REGION Network 15: DB62.DBX7.6 = Soot System Opacity
   // Word 4 bit 14
   RUNG wire#powerrail
      I_Contact( "10 DI_DATA".E700_OPACITY )
      { S7_Templates := "SrcType := Int" } GE_Contact(in1 := "100_BC_AUTO_SEQ_DB".CRNT_STEP, in2 := 240)
      Coil( %DB62.DBX7.6 )
   END_RUNG
   // the same network as SCL:
   %DB62.DBX7.6 := NOT "10 DI_DATA".E700_OPACITY AND ("100_BC_AUTO_SEQ_DB".CRNT_STEP >= 240);
END_REGION

REGION Network 16: DB62.DBX7.7 = Soot System Out of Range
   // Word 4 bit 15
   RUNG wire#powerrail
      "IDB_E700 Alarms"(Value := "12_AI_Data".E700SootContentIn, "Raw Value" := "IG Soot Content", Enable := true, "SHORT CIRCUIT VALUE" := 32000.0, "BROKEN WIRE VALUE" := -32000.0, "VERY LOW LEVEL VALUE (LL)" :=, "LOW LEVEL VALUE (L)" :=, "HIGH LEVEL VALUE (H)" :=, "VERY HIGH LEVEL VALUE (HH)" :=, OFFSET :=, "ALARM DELAY" :=, "Peak Value Reset" :=, "ALARM HH" =>, "ALARM H" =>, "ALARM L" =>, "ALARM LL" =>, "ALARM READING" => %DB62.DBX7.7, "Peak Value" =>, Alarm =>, Alarm_INT =>, "Enable Delay Time" :=, "High Value Release" :=)
   END_RUNG
   // the same network as SCL:
   "IDB_E700 Alarms"(Value := "12_AI_Data".E700SootContentIn,   // "502_ALM_ANALOG"
                     "Raw Value" := "IG Soot Content",
                     Enable := true,
                     "SHORT CIRCUIT VALUE" := 32000.0,
                     "BROKEN WIRE VALUE" := -32000.0,
                     "ALARM READING" => %DB62.DBX7.7);
END_REGION

REGION Network 17: DB62.DBX4.6 = E131 I&A Compresor Warning
   // Word 3 bit 6
   RUNG wire#powerrail
      I_Contact( "10 DI_DATA".E131_WRNG )
      Coil( %DB62.DBX4.6 )
   END_RUNG
   // the same network as SCL:
   %DB62.DBX4.6 := NOT "10 DI_DATA".E131_WRNG;
END_REGION

REGION Network 18: DB62.DBX4.7 = E131 I&A Compresor Not Running
   // Word 3 bit 7          Supresed. Not Available on The Bordeira
   RUNG wire#powerrail
      I_Contact( "10 DI_DATA".E131_OK )
      { S7_Templates := "SrcType := Int" } GT_Contact(in1 := "100_BC_AUTO_SEQ_DB".CRNT_STEP, in2 := 1)
      Contact( "AlwaysFALSE" )
      Coil( %DB62.DBX4.7 )
   END_RUNG
   // the same network as SCL:
   %DB62.DBX4.7 := NOT "10 DI_DATA".E131_OK AND ("100_BC_AUTO_SEQ_DB".CRNT_STEP > 1) AND "AlwaysFALSE";
END_REGION

REGION Network 19: DB62.DBX_ =IW98 - Flame Signal (FD-001)
   // Word 1 bit 12
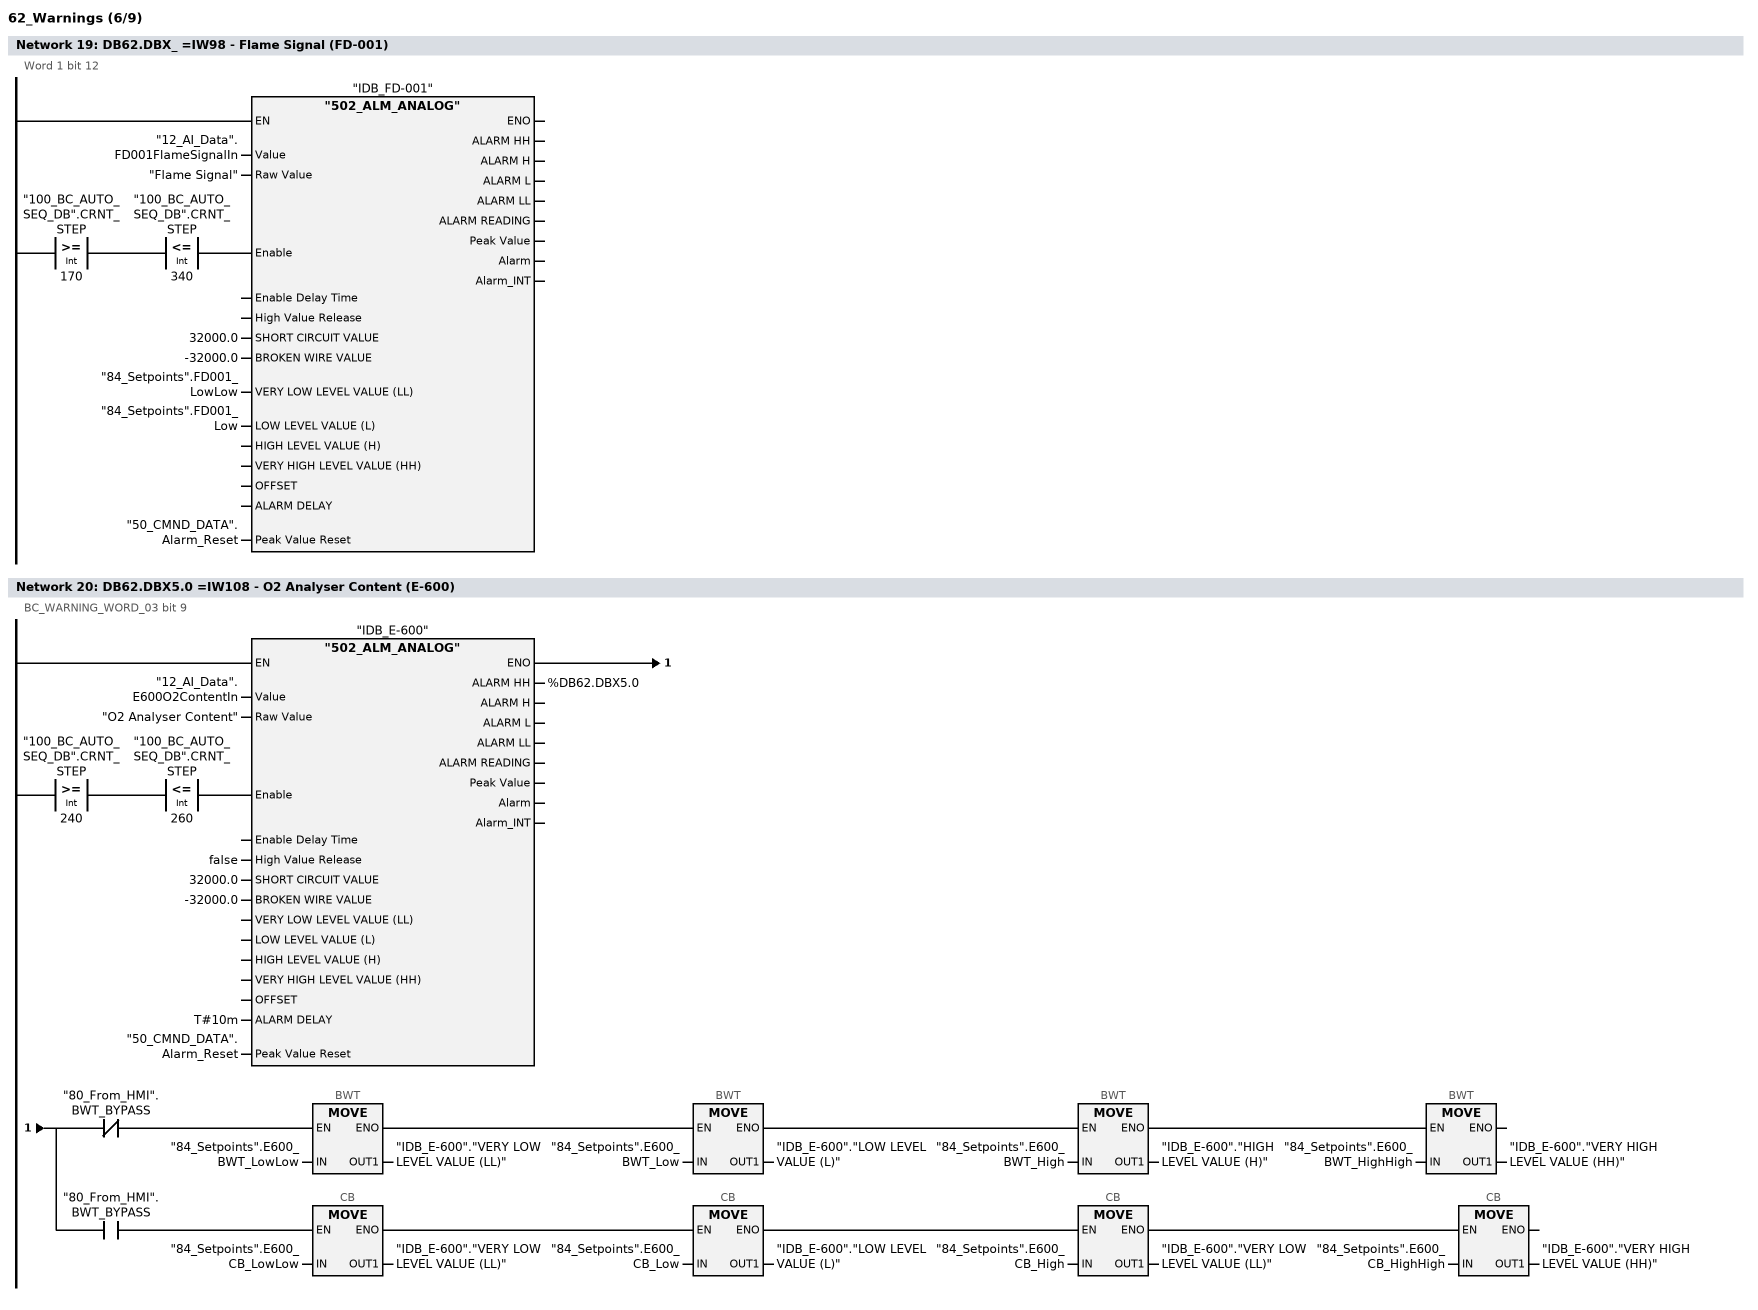
   RUNG wire#powerrail
      "IDB_FD-001"(Enable := wire#w1, Value := "12_AI_Data".FD001FlameSignalIn, "Raw Value" := "Flame Signal", "SHORT CIRCUIT VALUE" := 32000.0, "BROKEN WIRE VALUE" := -32000.0, "VERY LOW LEVEL VALUE (LL)" := "84_Setpoints".FD001_LowLow, "LOW LEVEL VALUE (L)" := "84_Setpoints".FD001_Low, "HIGH LEVEL VALUE (H)" :=, "VERY HIGH LEVEL VALUE (HH)" :=, OFFSET :=, "ALARM DELAY" :=, "Peak Value Reset" := "50_CMND_DATA".Alarm_Reset, "ALARM HH" =>, "ALARM H" =>, "ALARM L" =>, "ALARM LL" =>, "ALARM READING" =>, "Peak Value" =>, Alarm =>, Alarm_INT =>, "Enable Delay Time" :=, "High Value Release" :=)
   END_RUNG
   RUNG wire#powerrail
      { S7_Templates := "SrcType := Int" } GE_Contact(in1 := "100_BC_AUTO_SEQ_DB".CRNT_STEP, in2 := 170)
      { S7_Templates := "SrcType := Int" } LE_Contact(in1 := "100_BC_AUTO_SEQ_DB".CRNT_STEP, in2 := 340)
   END_RUNG wire#w1
   // the same network as SCL:
   "IDB_FD-001"(Value := "12_AI_Data".FD001FlameSignalIn,   // "502_ALM_ANALOG"
                "Raw Value" := "Flame Signal",
                Enable := ("100_BC_AUTO_SEQ_DB".CRNT_STEP >= 170) AND ("100_BC_AUTO_SEQ_DB".CRNT_STEP <= 340),
                "SHORT CIRCUIT VALUE" := 32000.0,
                "BROKEN WIRE VALUE" := -32000.0,
                "VERY LOW LEVEL VALUE (LL)" := "84_Setpoints".FD001_LowLow,
                "LOW LEVEL VALUE (L)" := "84_Setpoints".FD001_Low,
                "Peak Value Reset" := "50_CMND_DATA".Alarm_Reset);
END_REGION

REGION Network 20: DB62.DBX5.0 =IW108 - O2 Analyser Content (E-600)
   // BC_WARNING_WORD_03 bit 9
   RUNG wire#powerrail
      "IDB_E-600"(Enable := wire#w1, Value := "12_AI_Data".E600O2ContentIn, "Raw Value" := "O2 Analyser Content", "Enable Delay Time" :=, "High Value Release" := false, "SHORT CIRCUIT VALUE" := 32000.0, "BROKEN WIRE VALUE" := -32000.0, "VERY LOW LEVEL VALUE (LL)" :=, "LOW LEVEL VALUE (L)" :=, "HIGH LEVEL VALUE (H)" :=, "VERY HIGH LEVEL VALUE (HH)" :=, OFFSET :=, "ALARM DELAY" := T#10m, "Peak Value Reset" := "50_CMND_DATA".Alarm_Reset, "ALARM HH" => %DB62.DBX5.0, "ALARM H" =>, "ALARM L" =>, "ALARM LL" =>, "ALARM READING" =>, "Peak Value" =>, Alarm =>, Alarm_INT =>)
      wire#w2
      I_Contact( "80_From_HMI".BWT_BYPASS )
      Move(in := "84_Setpoints".E600_BWT_LowLow, out1 => "IDB_E-600"."VERY LOW LEVEL VALUE (LL)")   // BWT
      Move(in := "84_Setpoints".E600_BWT_Low, out1 => "IDB_E-600"."LOW LEVEL VALUE (L)")   // BWT
      Move(in := "84_Setpoints".E600_BWT_High, out1 => "IDB_E-600"."HIGH LEVEL VALUE (H)")   // BWT
      Move(in := "84_Setpoints".E600_BWT_HighHigh, out1 => "IDB_E-600"."VERY HIGH LEVEL VALUE (HH)")   // BWT
   END_RUNG
   RUNG wire#powerrail
      { S7_Templates := "SrcType := Int" } GE_Contact(in1 := "100_BC_AUTO_SEQ_DB".CRNT_STEP, in2 := 240)
      { S7_Templates := "SrcType := Int" } LE_Contact(in1 := "100_BC_AUTO_SEQ_DB".CRNT_STEP, in2 := 260)
   END_RUNG wire#w1
   RUNG wire#w2
      Contact( "80_From_HMI".BWT_BYPASS )
      Move(in := "84_Setpoints".E600_CB_LowLow, out1 => "IDB_E-600"."VERY LOW LEVEL VALUE (LL)")   // CB
      Move(in := "84_Setpoints".E600_CB_Low, out1 => "IDB_E-600"."LOW LEVEL VALUE (L)")   // CB
      Move(in := "84_Setpoints".E600_CB_High, out1 => "IDB_E-600"."VERY LOW LEVEL VALUE (LL)")   // CB
      Move(in := "84_Setpoints".E600_CB_HighHigh, out1 => "IDB_E-600"."VERY HIGH LEVEL VALUE (HH)")   // CB
   END_RUNG
   // the same network as SCL:
   "IDB_E-600"(Value := "12_AI_Data".E600O2ContentIn,   // "502_ALM_ANALOG"
               "Raw Value" := "O2 Analyser Content",
               Enable := ("100_BC_AUTO_SEQ_DB".CRNT_STEP >= 240) AND ("100_BC_AUTO_SEQ_DB".CRNT_STEP <= 260),
               "High Value Release" := false,
               "SHORT CIRCUIT VALUE" := 32000.0,
               "BROKEN WIRE VALUE" := -32000.0,
               "ALARM DELAY" := T#10m,
               "Peak Value Reset" := "50_CMND_DATA".Alarm_Reset,
               "ALARM HH" => %DB62.DBX5.0,
               ENO => #_w1);
   IF #_w1 AND NOT "80_From_HMI".BWT_BYPASS THEN
       "IDB_E-600"."VERY LOW LEVEL VALUE (LL)" := "84_Setpoints".E600_BWT_LowLow;   // BWT
       "IDB_E-600"."LOW LEVEL VALUE (L)" := "84_Setpoints".E600_BWT_Low;   // BWT
       "IDB_E-600"."HIGH LEVEL VALUE (H)" := "84_Setpoints".E600_BWT_High;   // BWT
       "IDB_E-600"."VERY HIGH LEVEL VALUE (HH)" := "84_Setpoints".E600_BWT_HighHigh;   // BWT
   END_IF;
   IF #_w1 AND "80_From_HMI".BWT_BYPASS THEN
       "IDB_E-600"."VERY LOW LEVEL VALUE (LL)" := "84_Setpoints".E600_CB_LowLow;   // CB
       "IDB_E-600"."LOW LEVEL VALUE (L)" := "84_Setpoints".E600_CB_Low;   // CB
       "IDB_E-600"."VERY LOW LEVEL VALUE (LL)" := "84_Setpoints".E600_CB_High;   // CB
       "IDB_E-600"."VERY HIGH LEVEL VALUE (HH)" := "84_Setpoints".E600_CB_HighHigh;   // CB
   END_IF;
END_REGION

REGION Network 21: DB62 DBX5.6 = Igniter Power Healthy
   // BC_WARNING_WORD_03_BIT_14
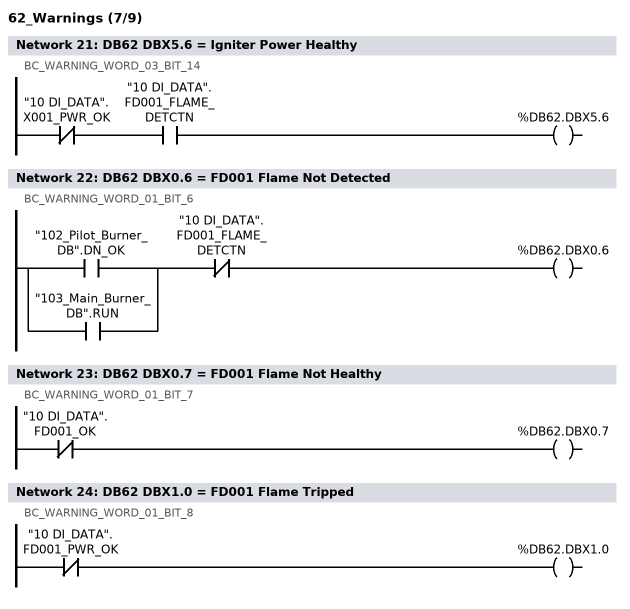
   RUNG wire#powerrail
      I_Contact( "10 DI_DATA".X001_PWR_OK )
      Contact( "10 DI_DATA".FD001_FLAME_DETCTN )
      Coil( %DB62.DBX5.6 )
   END_RUNG
   // the same network as SCL:
   %DB62.DBX5.6 := NOT "10 DI_DATA".X001_PWR_OK AND "10 DI_DATA".FD001_FLAME_DETCTN;
END_REGION

REGION Network 22: DB62 DBX0.6 = FD001 Flame Not Detected
   // BC_WARNING_WORD_01_BIT_6
   RUNG wire#powerrail
      Contact( "102_Pilot_Burner_DB".DN_OK )
      wire#w1
      I_Contact( "10 DI_DATA".FD001_FLAME_DETCTN )
      Coil( %DB62.DBX0.6 )
   END_RUNG
   RUNG wire#powerrail
      Contact( "103_Main_Burner_DB".RUN )
   END_RUNG wire#w1
   // the same network as SCL:
   %DB62.DBX0.6 := ("102_Pilot_Burner_DB".DN_OK OR "103_Main_Burner_DB".RUN) AND NOT "10 DI_DATA".FD001_FLAME_DETCTN;
END_REGION

REGION Network 23: DB62 DBX0.7 = FD001 Flame Not Healthy
   // BC_WARNING_WORD_01_BIT_7
   RUNG wire#powerrail
      I_Contact( "10 DI_DATA".FD001_OK )
      Coil( %DB62.DBX0.7 )
   END_RUNG
   // the same network as SCL:
   %DB62.DBX0.7 := NOT "10 DI_DATA".FD001_OK;
END_REGION

REGION Network 24: DB62 DBX1.0 = FD001 Flame Tripped
   // BC_WARNING_WORD_01_BIT_8
   RUNG wire#powerrail
      I_Contact( "10 DI_DATA".FD001_PWR_OK )
      Coil( %DB62.DBX1.0 )
   END_RUNG
   // the same network as SCL:
   %DB62.DBX1.0 := NOT "10 DI_DATA".FD001_PWR_OK;
END_REGION

REGION Network 25: Warning present
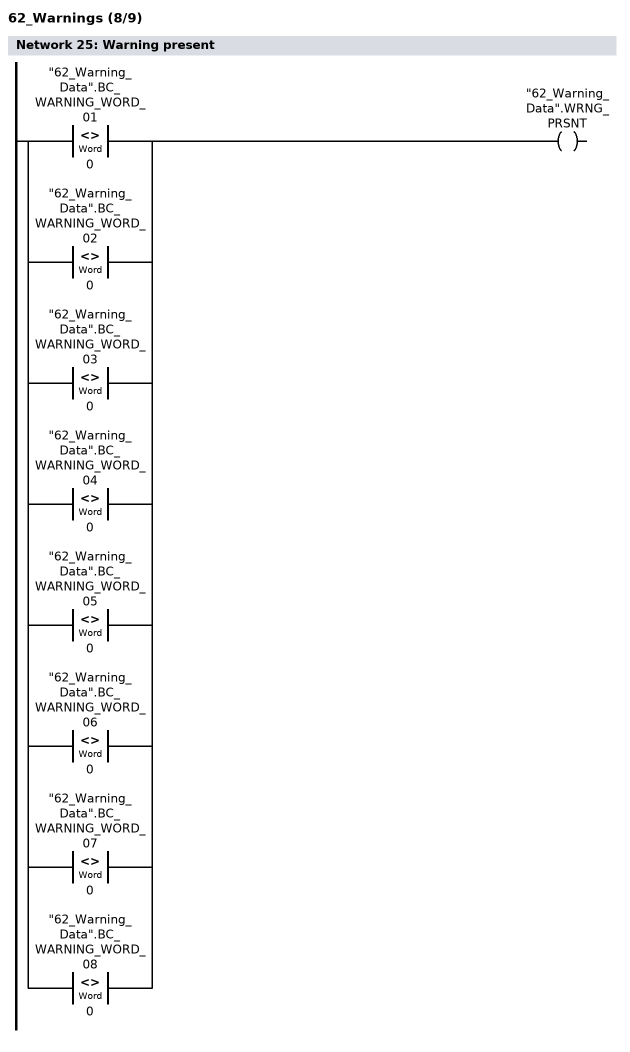
   RUNG wire#powerrail
      { S7_Templates := "SrcType := Word" } NE_Contact(in1 := "62_Warning_Data".BC_WARNING_WORD_01, in2 := 0)
      wire#w1
      Coil( "62_Warning_Data".WRNG_PRSNT )
   END_RUNG
   RUNG wire#powerrail
      { S7_Templates := "SrcType := Word" } NE_Contact(in1 := "62_Warning_Data".BC_WARNING_WORD_02, in2 := 0)
   END_RUNG wire#w1
   RUNG wire#powerrail
      { S7_Templates := "SrcType := Word" } NE_Contact(in1 := "62_Warning_Data".BC_WARNING_WORD_03, in2 := 0)
   END_RUNG wire#w1
   RUNG wire#powerrail
      { S7_Templates := "SrcType := Word" } NE_Contact(in1 := "62_Warning_Data".BC_WARNING_WORD_04, in2 := 0)
   END_RUNG wire#w1
   RUNG wire#powerrail
      { S7_Templates := "SrcType := Word" } NE_Contact(in1 := "62_Warning_Data".BC_WARNING_WORD_05, in2 := 0)
   END_RUNG wire#w1
   RUNG wire#powerrail
      { S7_Templates := "SrcType := Word" } NE_Contact(in1 := "62_Warning_Data".BC_WARNING_WORD_06, in2 := 0)
   END_RUNG wire#w1
   RUNG wire#powerrail
      { S7_Templates := "SrcType := Word" } NE_Contact(in1 := "62_Warning_Data".BC_WARNING_WORD_07, in2 := 0)
   END_RUNG wire#w1
   RUNG wire#powerrail
      { S7_Templates := "SrcType := Word" } NE_Contact(in1 := "62_Warning_Data".BC_WARNING_WORD_08, in2 := 0)
   END_RUNG wire#w1
   // the same network as SCL:
   "62_Warning_Data".WRNG_PRSNT := ("62_Warning_Data".BC_WARNING_WORD_01 <> 0) OR ("62_Warning_Data".BC_WARNING_WORD_02 <> 0) OR ("62_Warning_Data".BC_WARNING_WORD_03 <> 0) OR ("62_Warning_Data".BC_WARNING_WORD_04 <> 0) OR ("62_Warning_Data".BC_WARNING_WORD_05 <> 0) OR ("62_Warning_Data".BC_WARNING_WORD_06 <> 0) OR ("62_Warning_Data".BC_WARNING_WORD_07 <> 0) OR ("62_Warning_Data".BC_WARNING_WORD_08 <> 0);
END_REGION

REGION Network 26: New Warning Check
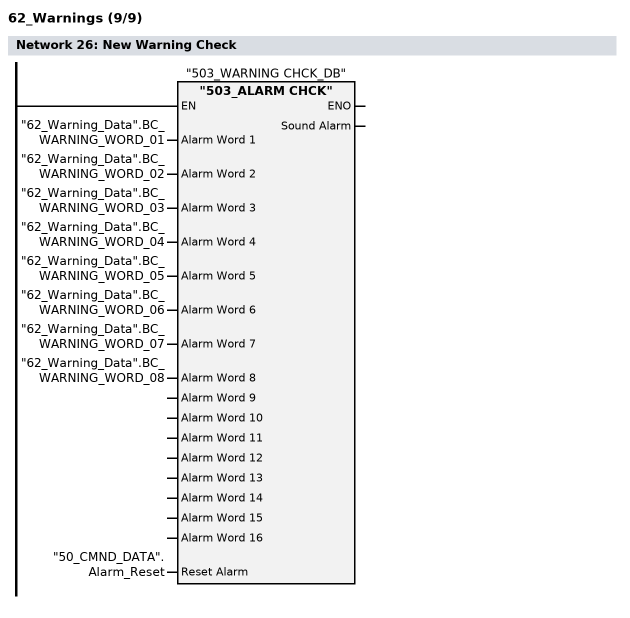
   RUNG wire#powerrail
      "503_WARNING CHCK_DB"("Alarm Word 1" := "62_Warning_Data".BC_WARNING_WORD_01, "Alarm Word 2" := "62_Warning_Data".BC_WARNING_WORD_02, "Alarm Word 3" := "62_Warning_Data".BC_WARNING_WORD_03, "Alarm Word 4" := "62_Warning_Data".BC_WARNING_WORD_04, "Alarm Word 5" := "62_Warning_Data".BC_WARNING_WORD_05, "Alarm Word 6" := "62_Warning_Data".BC_WARNING_WORD_06, "Alarm Word 7" := "62_Warning_Data".BC_WARNING_WORD_07, "Alarm Word 8" := "62_Warning_Data".BC_WARNING_WORD_08, "Alarm Word 9" :=, "Alarm Word 10" :=, "Alarm Word 11" :=, "Alarm Word 12" :=, "Alarm Word 13" :=, "Alarm Word 14" :=, "Alarm Word 15" :=, "Alarm Word 16" :=, "Reset Alarm" := "50_CMND_DATA".Alarm_Reset, "Sound Alarm" =>)
   END_RUNG
   // the same network as SCL:
   "503_WARNING CHCK_DB"("Alarm Word 1" := "62_Warning_Data".BC_WARNING_WORD_01,   // "503_ALARM CHCK"
                         "Alarm Word 2" := "62_Warning_Data".BC_WARNING_WORD_02,
                         "Alarm Word 3" := "62_Warning_Data".BC_WARNING_WORD_03,
                         "Alarm Word 4" := "62_Warning_Data".BC_WARNING_WORD_04,
                         "Alarm Word 5" := "62_Warning_Data".BC_WARNING_WORD_05,
                         "Alarm Word 6" := "62_Warning_Data".BC_WARNING_WORD_06,
                         "Alarm Word 7" := "62_Warning_Data".BC_WARNING_WORD_07,
                         "Alarm Word 8" := "62_Warning_Data".BC_WARNING_WORD_08,
                         "Reset Alarm" := "50_CMND_DATA".Alarm_Reset);
END_REGION
END_FUNCTION

FUNCTION "68_Sys_Status" : Void   // FC68, LAD
TITLE = System Status
{ S7_Optimized_Access := 'TRUE' }
AUTHOR : JRS
VERSION : 0.1
// For the determination of specific system status information as required by the code
   VAR_TEMP   // added for the SCL form of the ladder/FBD networks
      _w1 : Bool;
      _w2 : Bool;
   END_VAR
BEGIN

REGION Network 1: Valves At Initial
   // All valves in initial state
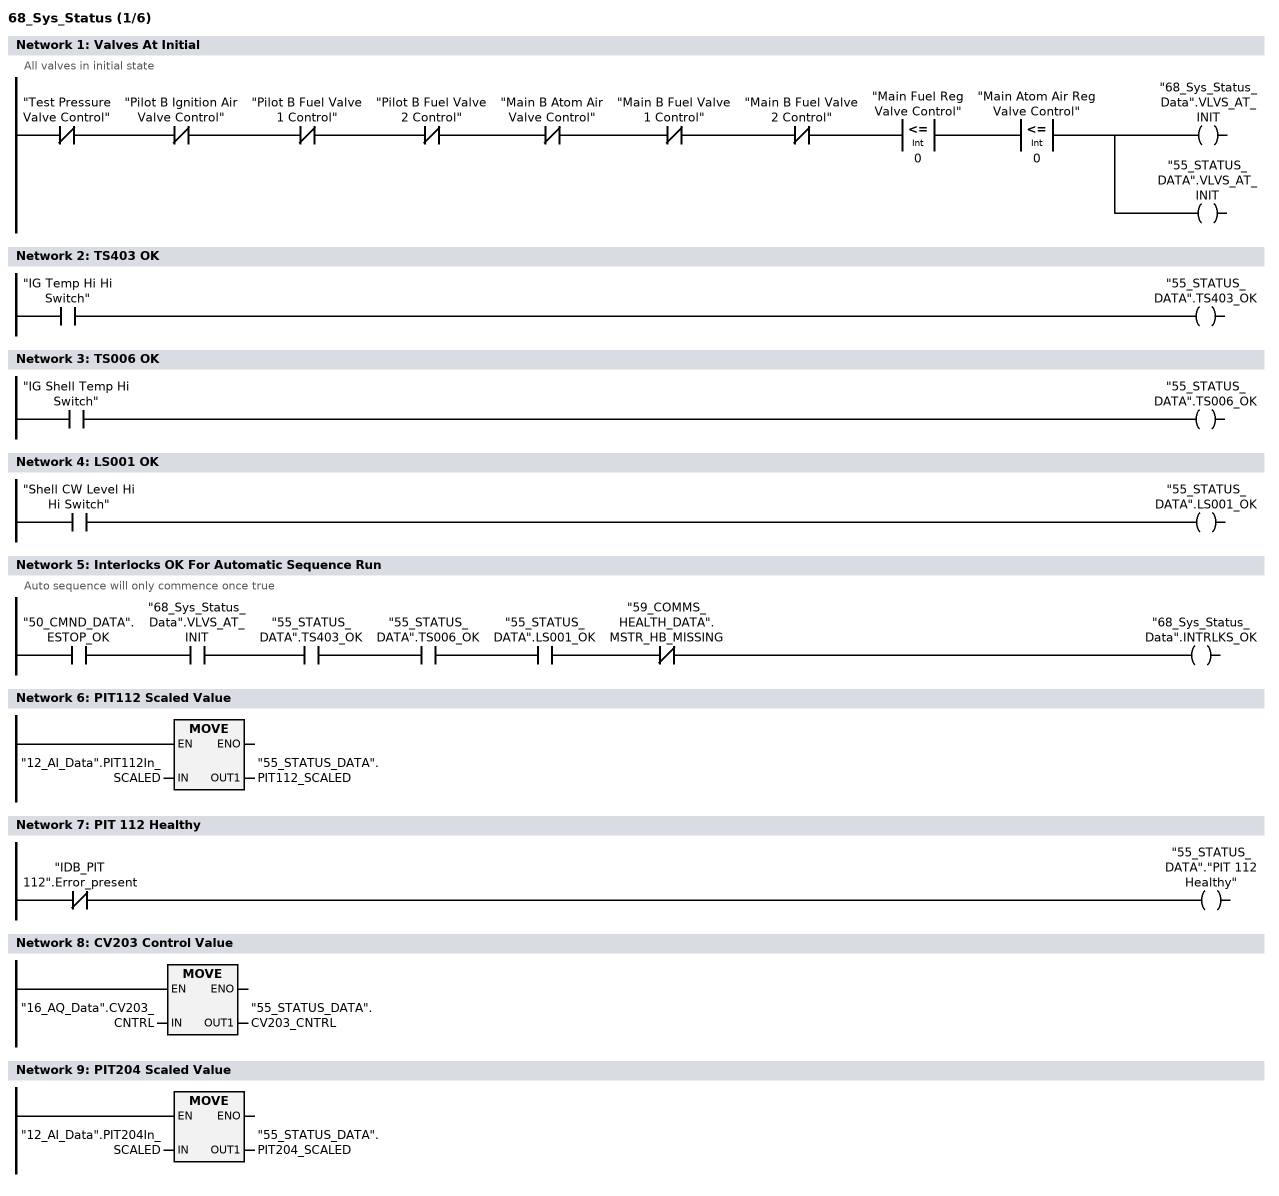
   RUNG wire#powerrail
      I_Contact( "Test Pressure Valve Control" )
      I_Contact( "Pilot B Ignition Air Valve Control" )
      I_Contact( "Pilot B Fuel Valve 1 Control" )
      I_Contact( "Pilot B Fuel Valve 2 Control" )
      I_Contact( "Main B Atom Air Valve Control" )
      I_Contact( "Main B Fuel Valve 1 Control" )
      I_Contact( "Main B Fuel Valve 2 Control" )
      { S7_Templates := "SrcType := Int" } LE_Contact(in1 := "Main Fuel Reg Valve Control", in2 := 0)
      { S7_Templates := "SrcType := Int" } LE_Contact(in1 := "Main Atom Air Reg Valve Control", in2 := 0)
      wire#w1
      Coil( "68_Sys_Status_Data".VLVS_AT_INIT )
   END_RUNG
   RUNG wire#w1
      Coil( "55_STATUS_DATA".VLVS_AT_INIT )
   END_RUNG
   // the same network as SCL:
   "68_Sys_Status_Data".VLVS_AT_INIT := NOT "Test Pressure Valve Control" AND NOT "Pilot B Ignition Air Valve Control" AND NOT "Pilot B Fuel Valve 1 Control" AND NOT "Pilot B Fuel Valve 2 Control" AND NOT "Main B Atom Air Valve Control" AND NOT "Main B Fuel Valve 1 Control" AND NOT "Main B Fuel Valve 2 Control" AND ("Main Fuel Reg Valve Control" <= 0) AND ("Main Atom Air Reg Valve Control" <= 0);
   "55_STATUS_DATA".VLVS_AT_INIT := "68_Sys_Status_Data".VLVS_AT_INIT;
END_REGION

REGION Network 2: TS403 OK
   RUNG wire#powerrail
      Contact( "IG Temp Hi Hi Switch" )
      Coil( "55_STATUS_DATA".TS403_OK )
   END_RUNG
   // the same network as SCL:
   "55_STATUS_DATA".TS403_OK := "IG Temp Hi Hi Switch";
END_REGION

REGION Network 3: TS006 OK
   RUNG wire#powerrail
      Contact( "IG Shell Temp Hi Switch" )
      Coil( "55_STATUS_DATA".TS006_OK )
   END_RUNG
   // the same network as SCL:
   "55_STATUS_DATA".TS006_OK := "IG Shell Temp Hi Switch";
END_REGION

REGION Network 4: LS001 OK
   RUNG wire#powerrail
      Contact( "Shell CW Level Hi Hi Switch" )
      Coil( "55_STATUS_DATA".LS001_OK )
   END_RUNG
   // the same network as SCL:
   "55_STATUS_DATA".LS001_OK := "Shell CW Level Hi Hi Switch";
END_REGION

REGION Network 5: Interlocks OK For Automatic Sequence Run
   // Auto sequence will only commence once true
   RUNG wire#powerrail
      Contact( "50_CMND_DATA".ESTOP_OK )
      Contact( "68_Sys_Status_Data".VLVS_AT_INIT )
      Contact( "55_STATUS_DATA".TS403_OK )
      Contact( "55_STATUS_DATA".TS006_OK )
      Contact( "55_STATUS_DATA".LS001_OK )
      I_Contact( "59_COMMS_HEALTH_DATA".MSTR_HB_MISSING )
      Coil( "68_Sys_Status_Data".INTRLKS_OK )
   END_RUNG
   // the same network as SCL:
   "68_Sys_Status_Data".INTRLKS_OK := "50_CMND_DATA".ESTOP_OK AND "68_Sys_Status_Data".VLVS_AT_INIT AND "55_STATUS_DATA".TS403_OK AND "55_STATUS_DATA".TS006_OK AND "55_STATUS_DATA".LS001_OK AND NOT "59_COMMS_HEALTH_DATA".MSTR_HB_MISSING;
END_REGION

REGION Network 6: PIT112 Scaled Value
   RUNG wire#powerrail
      Move(in := "12_AI_Data".PIT112In_SCALED, out1 => "55_STATUS_DATA".PIT112_SCALED)
   END_RUNG
   // the same network as SCL:
   "55_STATUS_DATA".PIT112_SCALED := "12_AI_Data".PIT112In_SCALED;
END_REGION

REGION Network 7: PIT 112 Healthy
   RUNG wire#powerrail
      I_Contact( "IDB_PIT 112".Error_present )
      Coil( "55_STATUS_DATA"."PIT 112 Healthy" )
   END_RUNG
   // the same network as SCL:
   "55_STATUS_DATA"."PIT 112 Healthy" := NOT "IDB_PIT 112".Error_present;
END_REGION

REGION Network 8: CV203 Control Value
   RUNG wire#powerrail
      Move(in := "16_AQ_Data".CV203_CNTRL, out1 => "55_STATUS_DATA".CV203_CNTRL)
   END_RUNG
   // the same network as SCL:
   "55_STATUS_DATA".CV203_CNTRL := "16_AQ_Data".CV203_CNTRL;
END_REGION

REGION Network 9: PIT204 Scaled Value
   RUNG wire#powerrail
      Move(in := "12_AI_Data".PIT204In_SCALED, out1 => "55_STATUS_DATA".PIT204_SCALED)
   END_RUNG
   // the same network as SCL:
   "55_STATUS_DATA".PIT204_SCALED := "12_AI_Data".PIT204In_SCALED;
END_REGION

REGION Network 10: P301 Enabled
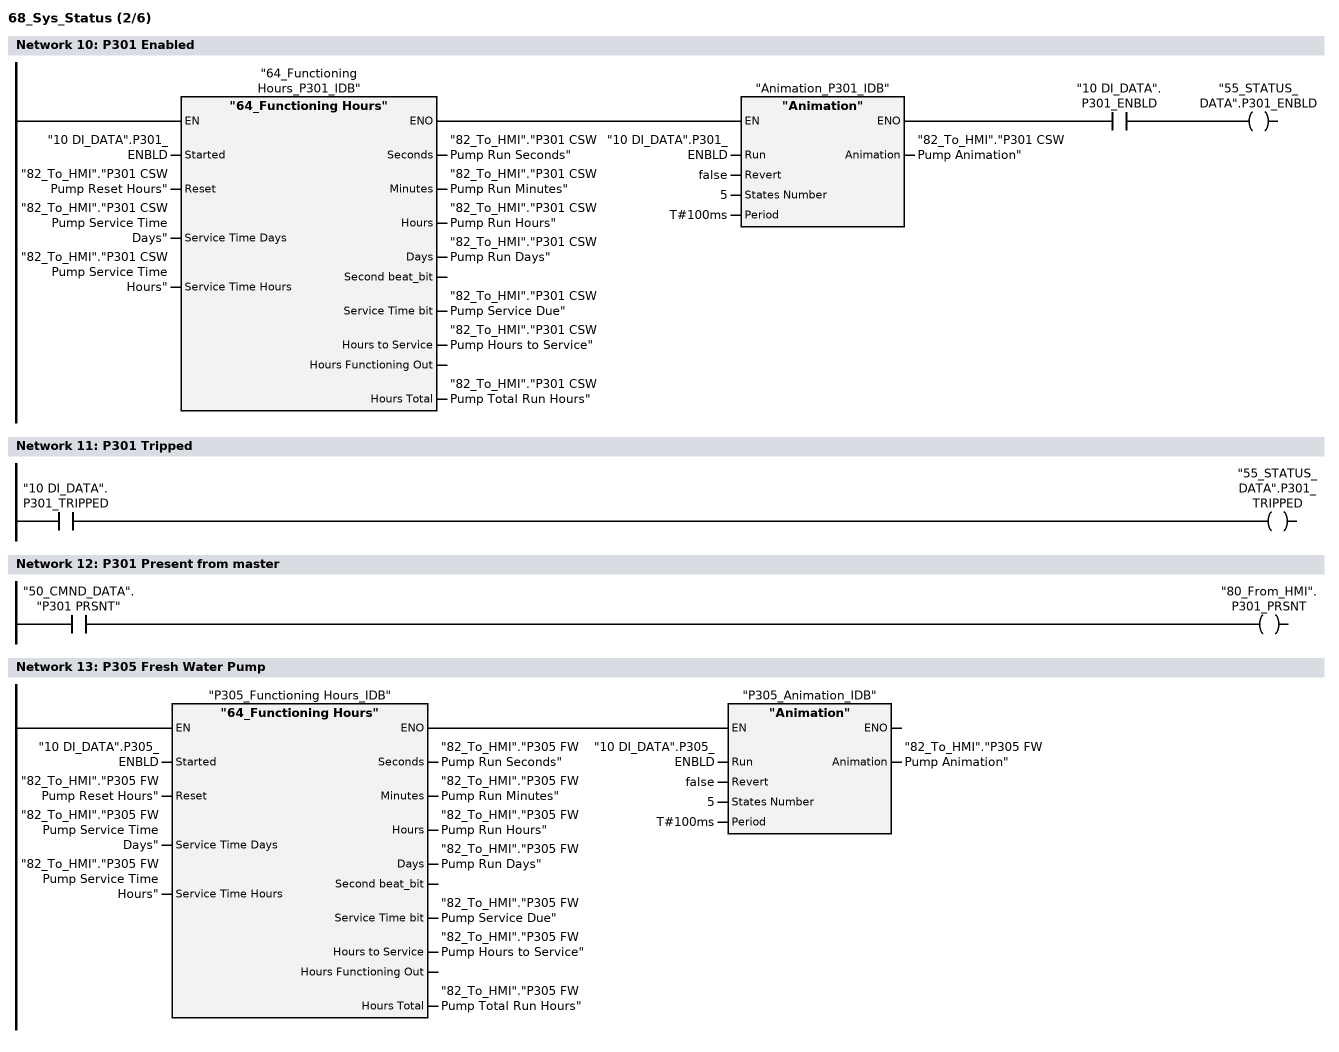
   RUNG wire#powerrail
      "64_Functioning Hours_P301_IDB"(Started := "10 DI_DATA".P301_ENBLD, Reset := "82_To_HMI"."P301 CSW Pump Reset Hours", "Service Time Days" := "82_To_HMI"."P301 CSW Pump Service Time Days", "Service Time Hours" := "82_To_HMI"."P301 CSW Pump Service Time Hours", Seconds => "82_To_HMI"."P301 CSW Pump Run Seconds", Minutes => "82_To_HMI"."P301 CSW Pump Run Minutes", Hours => "82_To_HMI"."P301 CSW Pump Run Hours", Days => "82_To_HMI"."P301 CSW Pump Run Days", "Second beat_bit" =>, "Service Time bit" => "82_To_HMI"."P301 CSW Pump Service Due", "Hours to Service" => "82_To_HMI"."P301 CSW Pump Hours to Service", "Hours Functioning Out" =>, "Hours Total" => "82_To_HMI"."P301 CSW Pump Total Run Hours")
      "Animation_P301_IDB"(Run := "10 DI_DATA".P301_ENBLD, Revert := false, "States Number" := 5, Period := T#100ms, Animation => "82_To_HMI"."P301 CSW Pump Animation")
      Contact( "10 DI_DATA".P301_ENBLD )
      Coil( "55_STATUS_DATA".P301_ENBLD )
   END_RUNG
   // the same network as SCL:
   "64_Functioning Hours_P301_IDB"(Started := "10 DI_DATA".P301_ENBLD,   // "64_Functioning Hours"
                           Reset := "82_To_HMI"."P301 CSW Pump Reset Hours",
                           "Service Time Days" := "82_To_HMI"."P301 CSW Pump Service Time Days",
                           "Service Time Hours" := "82_To_HMI"."P301 CSW Pump Service Time Hours",
                           Seconds => "82_To_HMI"."P301 CSW Pump Run Seconds",
                           Minutes => "82_To_HMI"."P301 CSW Pump Run Minutes",
                           Hours => "82_To_HMI"."P301 CSW Pump Run Hours",
                           Days => "82_To_HMI"."P301 CSW Pump Run Days",
                           "Service Time bit" => "82_To_HMI"."P301 CSW Pump Service Due",
                           "Hours to Service" => "82_To_HMI"."P301 CSW Pump Hours to Service",
                           "Hours Total" => "82_To_HMI"."P301 CSW Pump Total Run Hours",
                           ENO => #_w1);
   "Animation_P301_IDB"(EN := #_w1,   // "Animation"
                        Run := "10 DI_DATA".P301_ENBLD,
                        Revert := false,
                        "States Number" := 5,
                        Period := T#100ms,
                        Animation => "82_To_HMI"."P301 CSW Pump Animation",
                        ENO => #_w2);
   "55_STATUS_DATA".P301_ENBLD := #_w2 AND "10 DI_DATA".P301_ENBLD;
END_REGION

REGION Network 11: P301 Tripped
   RUNG wire#powerrail
      Contact( "10 DI_DATA".P301_TRIPPED )
      Coil( "55_STATUS_DATA".P301_TRIPPED )
   END_RUNG
   // the same network as SCL:
   "55_STATUS_DATA".P301_TRIPPED := "10 DI_DATA".P301_TRIPPED;
END_REGION

REGION Network 12: P301 Present from master
   RUNG wire#powerrail
      Contact( "50_CMND_DATA"."P301 PRSNT" )
      Coil( "80_From_HMI".P301_PRSNT )
   END_RUNG
   // the same network as SCL:
   "80_From_HMI".P301_PRSNT := "50_CMND_DATA"."P301 PRSNT";
END_REGION

REGION Network 13: P305 Fresh Water Pump
   RUNG wire#powerrail
      "P305_Functioning Hours_IDB"(Started := "10 DI_DATA".P305_ENBLD, Reset := "82_To_HMI"."P305 FW Pump Reset Hours", "Service Time Days" := "82_To_HMI"."P305 FW Pump Service Time Days", "Service Time Hours" := "82_To_HMI"."P305 FW Pump Service Time Hours", Seconds => "82_To_HMI"."P305 FW Pump Run Seconds", Minutes => "82_To_HMI"."P305 FW Pump Run Minutes", Hours => "82_To_HMI"."P305 FW Pump Run Hours", Days => "82_To_HMI"."P305 FW Pump Run Days", "Second beat_bit" =>, "Service Time bit" => "82_To_HMI"."P305 FW Pump Service Due", "Hours to Service" => "82_To_HMI"."P305 FW Pump Hours to Service", "Hours Functioning Out" =>, "Hours Total" => "82_To_HMI"."P305 FW Pump Total Run Hours")
      "P305_Animation_IDB"(Run := "10 DI_DATA".P305_ENBLD, Revert := false, "States Number" := 5, Period := T#100ms, Animation => "82_To_HMI"."P305 FW Pump Animation")
   END_RUNG
   // the same network as SCL:
   "P305_Functioning Hours_IDB"(Started := "10 DI_DATA".P305_ENBLD,   // "64_Functioning Hours"
                           Reset := "82_To_HMI"."P305 FW Pump Reset Hours",
                           "Service Time Days" := "82_To_HMI"."P305 FW Pump Service Time Days",
                           "Service Time Hours" := "82_To_HMI"."P305 FW Pump Service Time Hours",
                           Seconds => "82_To_HMI"."P305 FW Pump Run Seconds",
                           Minutes => "82_To_HMI"."P305 FW Pump Run Minutes",
                           Hours => "82_To_HMI"."P305 FW Pump Run Hours",
                           Days => "82_To_HMI"."P305 FW Pump Run Days",
                           "Service Time bit" => "82_To_HMI"."P305 FW Pump Service Due",
                           "Hours to Service" => "82_To_HMI"."P305 FW Pump Hours to Service",
                           "Hours Total" => "82_To_HMI"."P305 FW Pump Total Run Hours",
                           ENO => #_w1);
   IF #_w1 THEN
       "P305_Animation_IDB"(Run := "10 DI_DATA".P305_ENBLD,   // "Animation"
                            Revert := false,
                            "States Number" := 5,
                            Period := T#100ms,
                            Animation => "82_To_HMI"."P305 FW Pump Animation");
   END_IF;
END_REGION

REGION Network 14: E131 Running
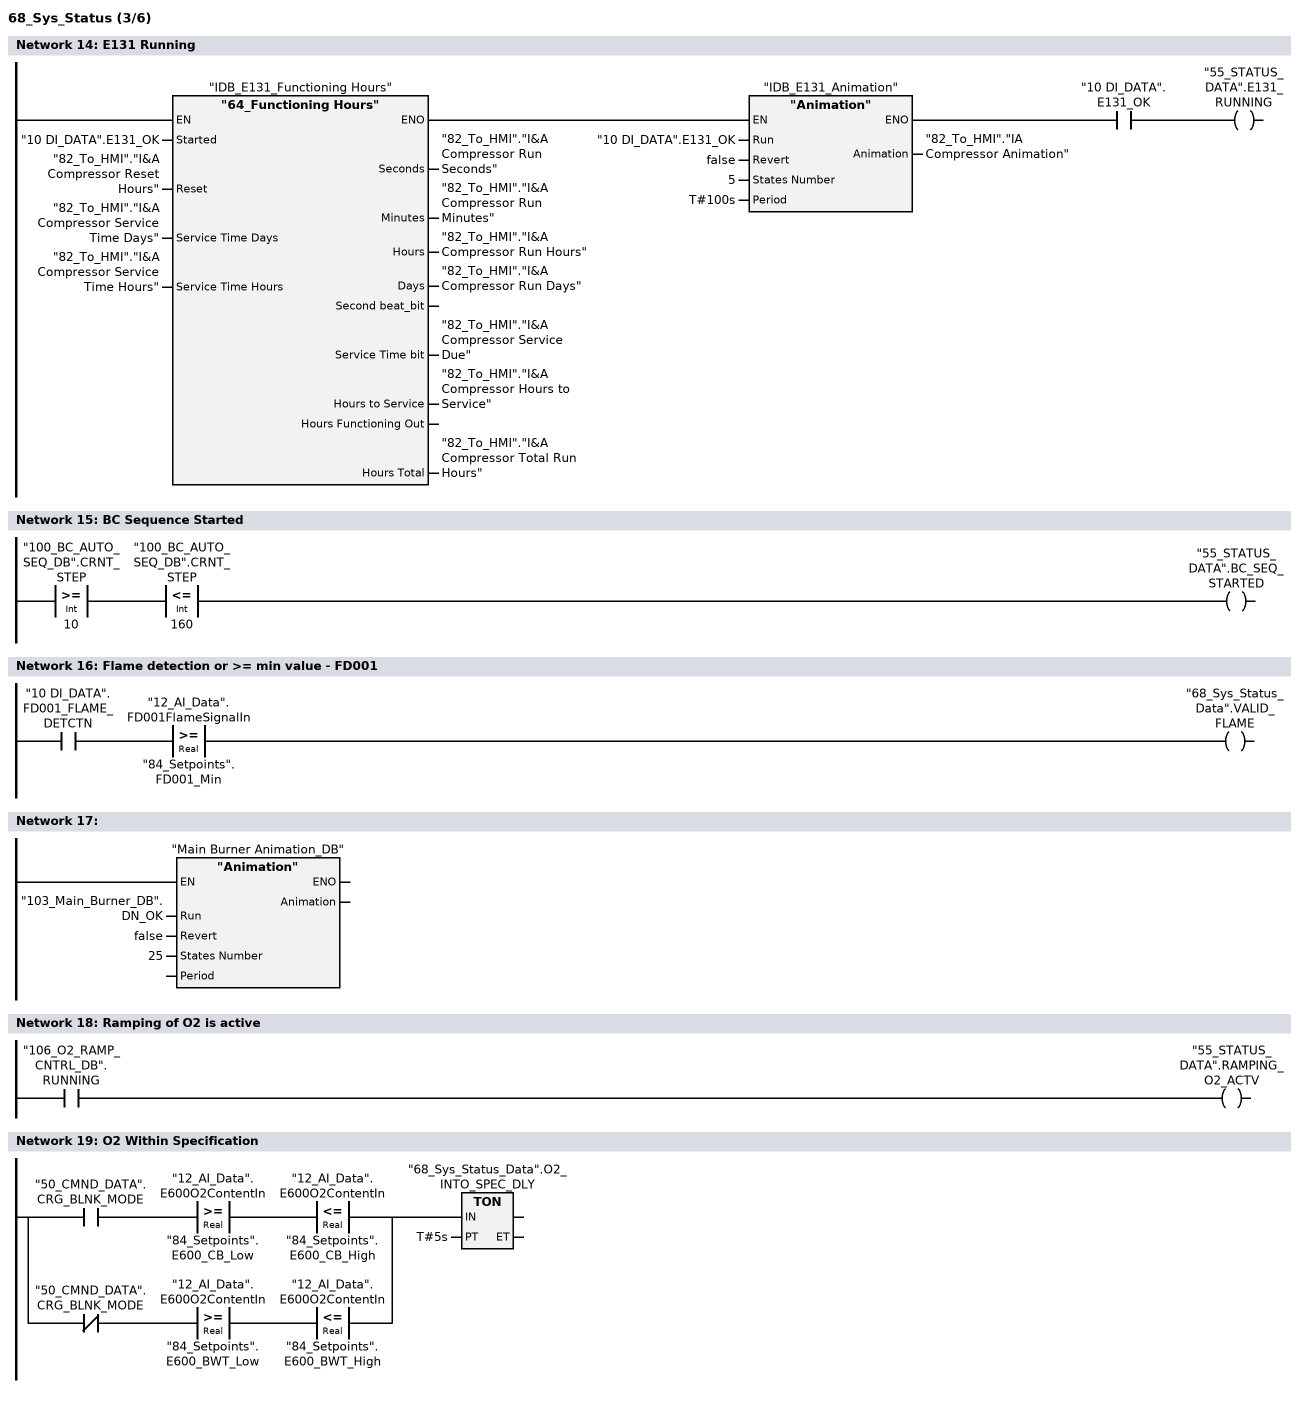
   RUNG wire#powerrail
      "IDB_E131_Functioning Hours"(Started := "10 DI_DATA".E131_OK, Reset := "82_To_HMI"."I&A Compressor Reset Hours", "Service Time Days" := "82_To_HMI"."I&A Compressor Service Time Days", "Service Time Hours" := "82_To_HMI"."I&A Compressor Service Time Hours", Seconds => "82_To_HMI"."I&A Compressor Run Seconds", Minutes => "82_To_HMI"."I&A Compressor Run Minutes", Hours => "82_To_HMI"."I&A Compressor Run Hours", Days => "82_To_HMI"."I&A Compressor Run Days", "Second beat_bit" =>, "Service Time bit" => "82_To_HMI"."I&A Compressor Service Due", "Hours to Service" => "82_To_HMI"."I&A Compressor Hours to Service", "Hours Functioning Out" =>, "Hours Total" => "82_To_HMI"."I&A Compressor Total Run Hours")
      "IDB_E131_Animation"(Run := "10 DI_DATA".E131_OK, Revert := false, "States Number" := 5, Period := T#100s, Animation => "82_To_HMI"."IA Compressor Animation")
      Contact( "10 DI_DATA".E131_OK )
      Coil( "55_STATUS_DATA".E131_RUNNING )
   END_RUNG
   // the same network as SCL:
   "IDB_E131_Functioning Hours"(Started := "10 DI_DATA".E131_OK,   // "64_Functioning Hours"
                           Reset := "82_To_HMI"."I&A Compressor Reset Hours",
                           "Service Time Days" := "82_To_HMI"."I&A Compressor Service Time Days",
                           "Service Time Hours" := "82_To_HMI"."I&A Compressor Service Time Hours",
                           Seconds => "82_To_HMI"."I&A Compressor Run Seconds",
                           Minutes => "82_To_HMI"."I&A Compressor Run Minutes",
                           Hours => "82_To_HMI"."I&A Compressor Run Hours",
                           Days => "82_To_HMI"."I&A Compressor Run Days",
                           "Service Time bit" => "82_To_HMI"."I&A Compressor Service Due",
                           "Hours to Service" => "82_To_HMI"."I&A Compressor Hours to Service",
                           "Hours Total" => "82_To_HMI"."I&A Compressor Total Run Hours",
                           ENO => #_w1);
   "IDB_E131_Animation"(EN := #_w1,   // "Animation"
                        Run := "10 DI_DATA".E131_OK,
                        Revert := false,
                        "States Number" := 5,
                        Period := T#100s,
                        Animation => "82_To_HMI"."IA Compressor Animation",
                        ENO => #_w2);
   "55_STATUS_DATA".E131_RUNNING := #_w2 AND "10 DI_DATA".E131_OK;
END_REGION

REGION Network 15: BC Sequence Started
   RUNG wire#powerrail
      { S7_Templates := "SrcType := Int" } GE_Contact(in1 := "100_BC_AUTO_SEQ_DB".CRNT_STEP, in2 := 10)
      { S7_Templates := "SrcType := Int" } LE_Contact(in1 := "100_BC_AUTO_SEQ_DB".CRNT_STEP, in2 := 160)
      Coil( "55_STATUS_DATA".BC_SEQ_STARTED )
   END_RUNG
   // the same network as SCL:
   "55_STATUS_DATA".BC_SEQ_STARTED := ("100_BC_AUTO_SEQ_DB".CRNT_STEP >= 10) AND ("100_BC_AUTO_SEQ_DB".CRNT_STEP <= 160);
END_REGION

REGION Network 16: Flame detection or >= min value - FD001
   RUNG wire#powerrail
      Contact( "10 DI_DATA".FD001_FLAME_DETCTN )
      { S7_Templates := "SrcType := Real" } GE_Contact(in1 := "12_AI_Data".FD001FlameSignalIn, in2 := "84_Setpoints".FD001_Min)
      Coil( "68_Sys_Status_Data".VALID_FLAME )
   END_RUNG
   // the same network as SCL:
   "68_Sys_Status_Data".VALID_FLAME := "10 DI_DATA".FD001_FLAME_DETCTN AND ("12_AI_Data".FD001FlameSignalIn >= "84_Setpoints".FD001_Min);
END_REGION

REGION Network 17
   RUNG wire#powerrail
      "Main Burner Animation_DB"(Run := "103_Main_Burner_DB".DN_OK, Revert := false, "States Number" := 25, Period :=, Animation =>)
   END_RUNG
   // the same network as SCL:
   "Main Burner Animation_DB"(Run := "103_Main_Burner_DB".DN_OK, Revert := false, "States Number" := 25);   // "Animation"
END_REGION

REGION Network 18: Ramping of O2 is active
   RUNG wire#powerrail
      Contact( "106_O2_RAMP_CNTRL_DB".RUNNING )
      Coil( "55_STATUS_DATA".RAMPING_O2_ACTV )
   END_RUNG
   // the same network as SCL:
   "55_STATUS_DATA".RAMPING_O2_ACTV := "106_O2_RAMP_CNTRL_DB".RUNNING;
END_REGION

REGION Network 19: O2 Within Specification
   "68_Sys_Status_Data".O2_INTO_SPEC_DLY.TON(IN := ("50_CMND_DATA".CRG_BLNK_MODE AND ("12_AI_Data".E600O2ContentIn >= "84_Setpoints".E600_CB_Low) AND ("12_AI_Data".E600O2ContentIn <= "84_Setpoints".E600_CB_High)) OR (NOT "50_CMND_DATA".CRG_BLNK_MODE AND ("12_AI_Data".E600O2ContentIn >= "84_Setpoints".E600_BWT_Low) AND ("12_AI_Data".E600O2ContentIn <= "84_Setpoints".E600_BWT_High)),
                           PT := T#5s);
END_REGION

REGION Network 20: O2 Within Specification
